// TIA Portal project "PolyMix_v0.1" (V14) (continued)
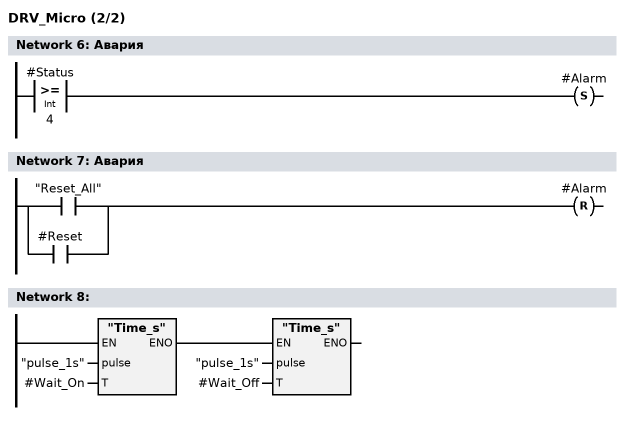
   RUNG wire#powerrail
      { S7_Templates := "SrcType := Int" } GE_Contact(in1 := #Status, in2 := 4)
      S_Coil( #Alarm )
   END_RUNG
   // the same network as SCL:
   IF #Status >= 4 THEN #Alarm := TRUE; END_IF;
END_REGION

REGION Network 7: Авария
   RUNG wire#powerrail
      Contact( "Reset_All" )
      wire#w1
      R_Coil( #Alarm )
   END_RUNG
   RUNG wire#powerrail
      Contact( #Reset )
   END_RUNG wire#w1
   // the same network as SCL:
   IF "Reset_All" OR #Reset THEN #Alarm := FALSE; END_IF;
END_REGION

REGION Network 8
   RUNG wire#powerrail
      "Time_s"(pulse := "pulse_1s", T := #Wait_On)
      "Time_s"(pulse := "pulse_1s", T := #Wait_Off)
   END_RUNG
   // the same network as SCL:
   "Time_s"(pulse := "pulse_1s", T := #Wait_On, ENO => #_w1);
   IF #_w1 THEN "Time_s"(pulse := "pulse_1s", T := #Wait_Off); END_IF;
END_REGION
END_FUNCTION_BLOCK

// folder: Modules

FUNCTION_BLOCK "DIx"   // FB200, LAD
{ S7_Optimized_Access := 'FALSE' }
VERSION : 0.1
// Input - входной сигнал контроллера
// pulse - частота фильтрации дребезга
// Signal - обработанный и отфильтрованный сигнал, используемый в дальнейшем
   VAR
      M1_FB_Ready : "DI_ex";   // I 0.0 - Мешалка 1 - готовность
      M1_FB_Run : "DI_ex";   // I 0.1 - Мешалка 1 - работа
      M2_FB_Ready : "DI_ex";   // I 0.2 - Мешалка 2 - готовность
      M2_FB_Run : "DI_ex";   // I 0.3 - Мешалка 2 - работа
      M3_FB_Ready : "DI_ex";   // I 0.4 - Мешалка 3 - готовность
      M3_FB_Run : "DI_ex";   // I 0.5 - Мешалка 3 - работа
      DD_FB_Ready : "DI_ex";   // I 0.6 - Дозатор сухого вещества - готовность
      Dos_FB_Run : "DI_ex";   // I 0.7 - Дозатор - работа
      DD_LLS : "DI_ex";   // I 1.0 - Дозатор сухого вещества - низкий уровень
      Vibro_FB_Ready : "DI_ex";   // I 1.1 - Вибратор - готовность
      Transporter : "DI_ex";   // I 1.2 - Пневмотранспортёр - готовность
      DL_FB_Ready : "DI_ex";   // I 1.3 - Дозатор жидкого вещества - готовность
      Dry_Run : "DI_ex";   // I 1.4 - Датчик протока
      AllBlock : "DI_ex";   // I 1.5 - Датчик перелива или Аварийная остановка
   END_VAR
   VAR_TEMP   // added for the SCL form of the ladder/FBD networks
      _w1 : Bool;
      _w2 : Bool;
   END_VAR
BEGIN

REGION Network 1: Мешалка 1
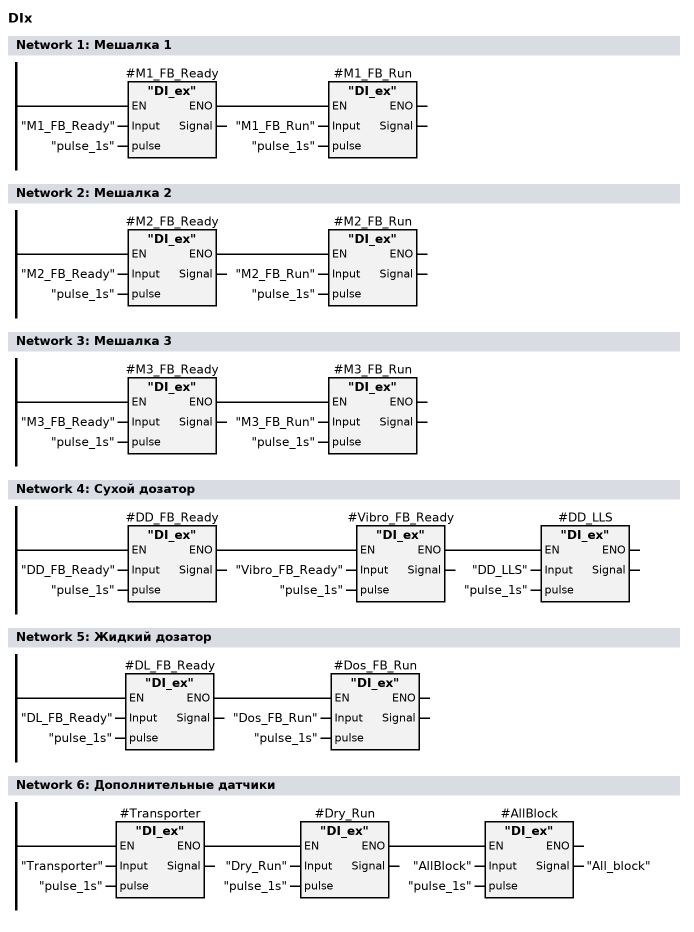
   RUNG wire#powerrail
      #M1_FB_Ready(Input := "M1_FB_Ready", pulse := "pulse_1s", Signal =>)
      #M1_FB_Run(Input := "M1_FB_Run", pulse := "pulse_1s", Signal =>)
   END_RUNG
   // the same network as SCL:
   #M1_FB_Ready(Input := "M1_FB_Ready", pulse := "pulse_1s", ENO => #_w1);   // "DI_ex"
   IF #_w1 THEN
       #M1_FB_Run(Input := "M1_FB_Run", pulse := "pulse_1s");   // "DI_ex"
   END_IF;
END_REGION

REGION Network 2: Мешалка 2
   RUNG wire#powerrail
      #M2_FB_Ready(Input := "M2_FB_Ready", pulse := "pulse_1s", Signal =>)
      #M2_FB_Run(Input := "M2_FB_Run", pulse := "pulse_1s", Signal =>)
   END_RUNG
   // the same network as SCL:
   #M2_FB_Ready(Input := "M2_FB_Ready", pulse := "pulse_1s", ENO => #_w1);   // "DI_ex"
   IF #_w1 THEN
       #M2_FB_Run(Input := "M2_FB_Run", pulse := "pulse_1s");   // "DI_ex"
   END_IF;
END_REGION

REGION Network 3: Мешалка 3
   RUNG wire#powerrail
      #M3_FB_Ready(Input := "M3_FB_Ready", pulse := "pulse_1s", Signal =>)
      #M3_FB_Run(Input := "M3_FB_Run", pulse := "pulse_1s", Signal =>)
   END_RUNG
   // the same network as SCL:
   #M3_FB_Ready(Input := "M3_FB_Ready", pulse := "pulse_1s", ENO => #_w1);   // "DI_ex"
   IF #_w1 THEN
       #M3_FB_Run(Input := "M3_FB_Run", pulse := "pulse_1s");   // "DI_ex"
   END_IF;
END_REGION

REGION Network 4: Сухой дозатор
   RUNG wire#powerrail
      #DD_FB_Ready(Input := "DD_FB_Ready", pulse := "pulse_1s", Signal =>)
      #Vibro_FB_Ready(Input := "Vibro_FB_Ready", pulse := "pulse_1s", Signal =>)
      #DD_LLS(Input := "DD_LLS", pulse := "pulse_1s", Signal =>)
   END_RUNG
   // the same network as SCL:
   #DD_FB_Ready(Input := "DD_FB_Ready", pulse := "pulse_1s", ENO => #_w1);   // "DI_ex"
   #Vibro_FB_Ready(EN := #_w1, Input := "Vibro_FB_Ready", pulse := "pulse_1s", ENO => #_w2);   // "DI_ex"
   IF #_w2 THEN
       #DD_LLS(Input := "DD_LLS", pulse := "pulse_1s");   // "DI_ex"
   END_IF;
END_REGION

REGION Network 5: Жидкий дозатор
   RUNG wire#powerrail
      #DL_FB_Ready(Input := "DL_FB_Ready", pulse := "pulse_1s", Signal =>)
      #Dos_FB_Run(Input := "Dos_FB_Run", pulse := "pulse_1s", Signal =>)
   END_RUNG
   // the same network as SCL:
   #DL_FB_Ready(Input := "DL_FB_Ready", pulse := "pulse_1s", ENO => #_w1);   // "DI_ex"
   IF #_w1 THEN
       #Dos_FB_Run(Input := "Dos_FB_Run", pulse := "pulse_1s");   // "DI_ex"
   END_IF;
END_REGION

REGION Network 6: Дополнительные датчики
   RUNG wire#powerrail
      #Transporter(Input := "Transporter", pulse := "pulse_1s", Signal =>)
      #Dry_Run(Input := "Dry_Run", pulse := "pulse_1s", Signal =>)
      #AllBlock(Input := "AllBlock", pulse := "pulse_1s", Signal => "All_block")
   END_RUNG
   // the same network as SCL:
   #Transporter(Input := "Transporter", pulse := "pulse_1s", ENO => #_w1);   // "DI_ex"
   #Dry_Run(EN := #_w1, Input := "Dry_Run", pulse := "pulse_1s", ENO => #_w2);   // "DI_ex"
   IF #_w2 THEN
       #AllBlock(Input := "AllBlock", pulse := "pulse_1s", Signal => "All_block");   // "DI_ex"
   END_IF;
END_REGION
END_FUNCTION_BLOCK

FUNCTION_BLOCK "DOx"   // FB201, LAD
{ S7_Optimized_Access := 'FALSE' }
VERSION : 0.1
// Start - управляющий сигнал из программы
// Q - выходной сигнал контроллера
// pulse - кратность времени в импульсном режиме
   VAR
      M1_CMD : "DO_ex";   // Q 0.0 - Мешалка 1 - запуск
      M2_CMD : "DO_ex";   // Q 0.1 - Мешалка 2 - запуск
      M3_CMD : "DO_ex";   // Q 0.2 - Мешалка 3 - запуск
      DD_CMD : "DO_ex";   // Q 0.3 - Дозатор сухого вещества - запуск
      Vibro_CMD : "DO_ex";   // Q 0.4 - Вибратор - запуск
      DL_CMD : "DO_ex";   // Q 0.5 - Дозатор жидкого вещества - запуск
      KC1_CMD : "DO_ex";   // Q 0.6 - Соленоидный клапан КС1
      LED_Dry_Run : "DO_ex";   // Q 0.7 - LED - сухой ход
      LED_Alarm : "DO_ex";   // Q 1.0 - LED - общая авария
      LED_Empty : "DO_ex";   // Q 1.1 - LED - бункер пуст
   END_VAR
   VAR_TEMP   // added for the SCL form of the ladder/FBD networks
      _w1 : Bool;
      _w2 : Bool;
   END_VAR
BEGIN

REGION Network 1: Мешалки 1-3
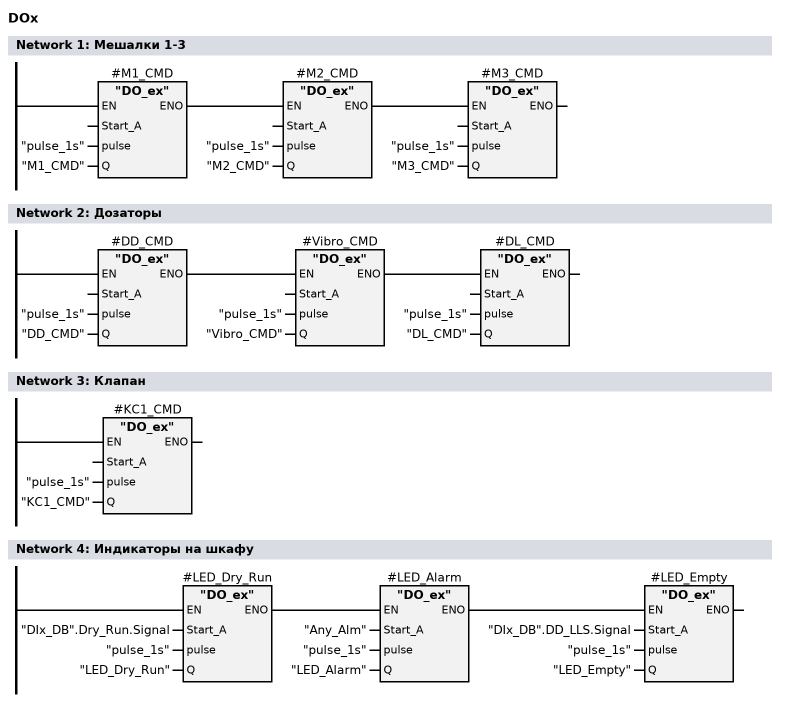
   RUNG wire#powerrail
      #M1_CMD(Start_A :=, pulse := "pulse_1s", Q := "M1_CMD")
      #M2_CMD(Start_A :=, pulse := "pulse_1s", Q := "M2_CMD")
      #M3_CMD(Start_A :=, pulse := "pulse_1s", Q := "M3_CMD")
   END_RUNG
   // the same network as SCL:
   #M1_CMD(pulse := "pulse_1s", Q := "M1_CMD", ENO => #_w1);   // "DO_ex"
   #M2_CMD(EN := #_w1, pulse := "pulse_1s", Q := "M2_CMD", ENO => #_w2);   // "DO_ex"
   IF #_w2 THEN
       #M3_CMD(pulse := "pulse_1s", Q := "M3_CMD");   // "DO_ex"
   END_IF;
END_REGION

REGION Network 2: Дозаторы
   RUNG wire#powerrail
      #DD_CMD(Start_A :=, pulse := "pulse_1s", Q := "DD_CMD")
      #Vibro_CMD(Start_A :=, pulse := "pulse_1s", Q := "Vibro_CMD")
      #DL_CMD(Start_A :=, pulse := "pulse_1s", Q := "DL_CMD")
   END_RUNG
   // the same network as SCL:
   #DD_CMD(pulse := "pulse_1s", Q := "DD_CMD", ENO => #_w1);   // "DO_ex"
   #Vibro_CMD(EN := #_w1, pulse := "pulse_1s", Q := "Vibro_CMD", ENO => #_w2);   // "DO_ex"
   IF #_w2 THEN
       #DL_CMD(pulse := "pulse_1s", Q := "DL_CMD");   // "DO_ex"
   END_IF;
END_REGION

REGION Network 3: Клапан
   RUNG wire#powerrail
      #KC1_CMD(Start_A :=, pulse := "pulse_1s", Q := "KC1_CMD")
   END_RUNG
   // the same network as SCL:
   #KC1_CMD(pulse := "pulse_1s", Q := "KC1_CMD");   // "DO_ex"
END_REGION

REGION Network 4: Индикаторы на шкафу
   RUNG wire#powerrail
      #LED_Dry_Run(Start_A := "DIx_DB".Dry_Run.Signal, pulse := "pulse_1s", Q := "LED_Dry_Run")
      #LED_Alarm(Start_A := "Any_Alm", pulse := "pulse_1s", Q := "LED_Alarm")
      #LED_Empty(Start_A := "DIx_DB".DD_LLS.Signal, pulse := "pulse_1s", Q := "LED_Empty")
   END_RUNG
   // the same network as SCL:
   #LED_Dry_Run(Start_A := "DIx_DB".Dry_Run.Signal, pulse := "pulse_1s", Q := "LED_Dry_Run", ENO => #_w1);   // "DO_ex"
   #LED_Alarm(EN := #_w1, Start_A := "Any_Alm", pulse := "pulse_1s", Q := "LED_Alarm", ENO => #_w2);   // "DO_ex"
   IF #_w2 THEN
       #LED_Empty(Start_A := "DIx_DB".DD_LLS.Signal, pulse := "pulse_1s", Q := "LED_Empty");   // "DO_ex"
   END_IF;
END_REGION
END_FUNCTION_BLOCK

FUNCTION_BLOCK "Micro"   // FB207, LAD
{ S7_Optimized_Access := 'FALSE' }
VERSION : 0.1
   VAR
      KC1 : "DRV_Micro";   // Соленоидный клапан
   END_VAR
   // KC1.No_FB := true;
BEGIN

REGION Network 1
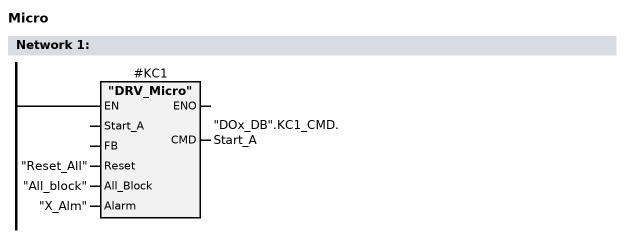
   RUNG wire#powerrail
      #KC1(Start_A :=, FB :=, Reset := "Reset_All", All_Block := "All_block", Alarm := "X_Alm", CMD => "DOx_DB".KC1_CMD.Start_A)
   END_RUNG
   // the same network as SCL:
   #KC1(Reset := "Reset_All", All_Block := "All_block", Alarm := "X_Alm", CMD => "DOx_DB".KC1_CMD.Start_A);   // "DRV_Micro"
END_REGION
END_FUNCTION_BLOCK

// folder: System

FUNCTION "DRV_pulse" : Void   // FC100, LAD
{ S7_Optimized_Access := 'FALSE' }
VERSION : 0.1
   VAR_TEMP   // added for the SCL form of the ladder/FBD networks
      _w1 : Bool;
      _w2 : Bool;
   END_VAR
BEGIN

REGION Network 1
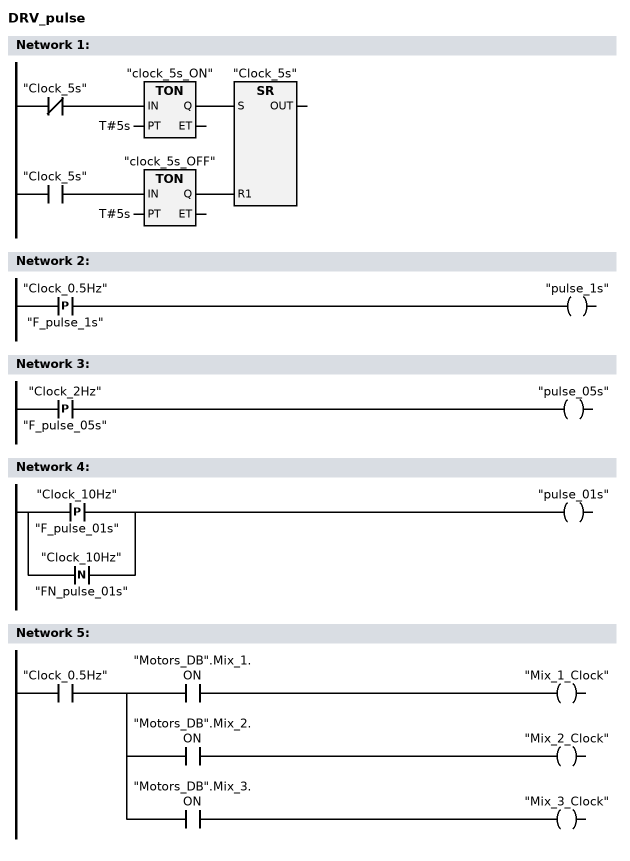
   "clock_5s_ON".TON(IN := NOT "Clock_5s", PT := T#5s);
   "clock_5s_OFF".TON(IN := "Clock_5s", PT := T#5s);
   IF "clock_5s_ON".Q THEN
       "Clock_5s" := TRUE;   // SR flip-flop
   END_IF;
   IF "clock_5s_OFF".Q THEN "Clock_5s" := FALSE; END_IF;
END_REGION

REGION Network 2
   RUNG wire#powerrail
      P_Contact(operand := "Clock_0.5Hz", bit := "F_pulse_1s")
      Coil( "pulse_1s" )
   END_RUNG
   // the same network as SCL:
   #_w1 := "Clock_0.5Hz" AND NOT "F_pulse_1s";   // rising edge of "Clock_0.5Hz"
   "F_pulse_1s" := "Clock_0.5Hz";
   "pulse_1s" := #_w1;
END_REGION

REGION Network 3
   RUNG wire#powerrail
      P_Contact(operand := "Clock_2Hz", bit := "F_pulse_05s")
      Coil( "pulse_05s" )
   END_RUNG
   // the same network as SCL:
   #_w1 := "Clock_2Hz" AND NOT "F_pulse_05s";   // rising edge of "Clock_2Hz"
   "F_pulse_05s" := "Clock_2Hz";
   "pulse_05s" := #_w1;
END_REGION

REGION Network 4
   RUNG wire#powerrail
      P_Contact(operand := "Clock_10Hz", bit := "F_pulse_01s")
      wire#w1
      Coil( "pulse_01s" )
   END_RUNG
   RUNG wire#powerrail
      N_Contact(operand := "Clock_10Hz", bit := "FN_pulse_01s")
   END_RUNG wire#w1
   // the same network as SCL:
   #_w1 := "Clock_10Hz" AND NOT "F_pulse_01s";   // rising edge of "Clock_10Hz"
   "F_pulse_01s" := "Clock_10Hz";
   #_w2 := NOT "Clock_10Hz" AND "FN_pulse_01s";   // falling edge of "Clock_10Hz"
   "FN_pulse_01s" := "Clock_10Hz";
   "pulse_01s" := #_w1 OR #_w2;
END_REGION

REGION Network 5
   RUNG wire#powerrail
      Contact( "Clock_0.5Hz" )
      wire#w1
      Contact( "Motors_DB".Mix_1.ON )
      Coil( "Mix_1_Clock" )
   END_RUNG
   RUNG wire#w1
      Contact( "Motors_DB".Mix_2.ON )
      Coil( "Mix_2_Clock" )
   END_RUNG
   RUNG wire#w1
      Contact( "Motors_DB".Mix_3.ON )
      Coil( "Mix_3_Clock" )
   END_RUNG
   // the same network as SCL:
   "Mix_1_Clock" := "Clock_0.5Hz" AND "Motors_DB".Mix_1.ON;
   "Mix_2_Clock" := "Clock_0.5Hz" AND "Motors_DB".Mix_2.ON;
   "Mix_3_Clock" := "Clock_0.5Hz" AND "Motors_DB".Mix_3.ON;
END_REGION
END_FUNCTION

FUNCTION "DRV_End" : Void   // FC101, LAD
{ S7_Optimized_Access := 'TRUE' }
VERSION : 0.1
BEGIN

REGION Network 1: Одно из устройств нижнего уровня в ручном режиме
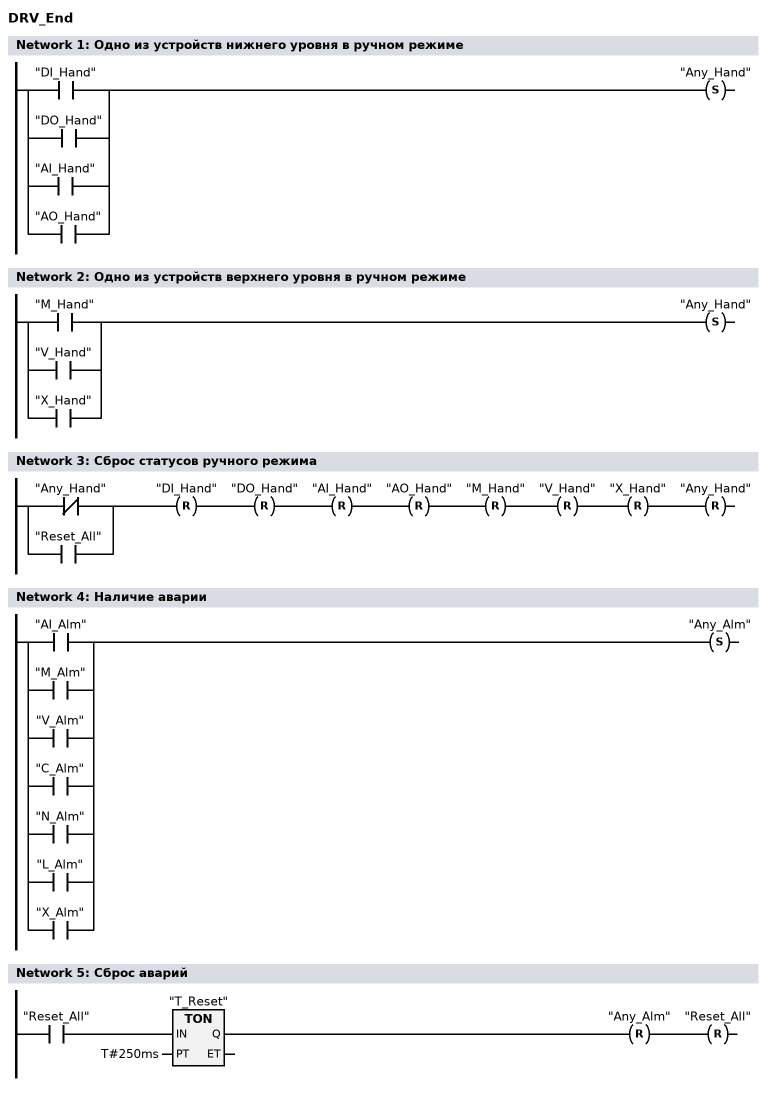
   RUNG wire#powerrail
      Contact( "DI_Hand" )
      wire#w1
      S_Coil( "Any_Hand" )
   END_RUNG
   RUNG wire#powerrail
      Contact( "DO_Hand" )
   END_RUNG wire#w1
   RUNG wire#powerrail
      Contact( "AI_Hand" )
   END_RUNG wire#w1
   RUNG wire#powerrail
      Contact( "AO_Hand" )
   END_RUNG wire#w1
   // the same network as SCL:
   IF "DI_Hand" OR "DO_Hand" OR "AI_Hand" OR "AO_Hand" THEN "Any_Hand" := TRUE; END_IF;
END_REGION

REGION Network 2: Одно из устройств верхнего уровня в ручном режиме
   RUNG wire#powerrail
      Contact( "M_Hand" )
      wire#w1
      S_Coil( "Any_Hand" )
   END_RUNG
   RUNG wire#powerrail
      Contact( "V_Hand" )
   END_RUNG wire#w1
   RUNG wire#powerrail
      Contact( "X_Hand" )
   END_RUNG wire#w1
   // the same network as SCL:
   IF "M_Hand" OR "V_Hand" OR "X_Hand" THEN "Any_Hand" := TRUE; END_IF;
END_REGION

REGION Network 3: Сброс статусов ручного режима
   RUNG wire#powerrail
      I_Contact( "Any_Hand" )
      wire#w1
      R_Coil( "DI_Hand" )
      R_Coil( "DO_Hand" )
      R_Coil( "AI_Hand" )
      R_Coil( "AO_Hand" )
      R_Coil( "M_Hand" )
      R_Coil( "V_Hand" )
      R_Coil( "X_Hand" )
      R_Coil( "Any_Hand" )
   END_RUNG
   RUNG wire#powerrail
      Contact( "Reset_All" )
   END_RUNG wire#w1
   // the same network as SCL:
   IF NOT "Any_Hand" OR "Reset_All" THEN
       "DI_Hand" := FALSE;
       "DO_Hand" := FALSE;
       "AI_Hand" := FALSE;
       "AO_Hand" := FALSE;
       "M_Hand" := FALSE;
       "V_Hand" := FALSE;
       "X_Hand" := FALSE;
       "Any_Hand" := FALSE;
   END_IF;
END_REGION

REGION Network 4: Наличие аварии
   RUNG wire#powerrail
      Contact( "AI_Alm" )
      wire#w1
      S_Coil( "Any_Alm" )
   END_RUNG
   RUNG wire#powerrail
      Contact( "M_Alm" )
   END_RUNG wire#w1
   RUNG wire#powerrail
      Contact( "V_Alm" )
   END_RUNG wire#w1
   RUNG wire#powerrail
      Contact( "C_Alm" )
   END_RUNG wire#w1
   RUNG wire#powerrail
      Contact( "N_Alm" )
   END_RUNG wire#w1
   RUNG wire#powerrail
      Contact( "L_Alm" )
   END_RUNG wire#w1
   RUNG wire#powerrail
      Contact( "X_Alm" )
   END_RUNG wire#w1
   // the same network as SCL:
   IF "AI_Alm" OR "M_Alm" OR "V_Alm" OR "C_Alm" OR "N_Alm" OR "L_Alm" OR "X_Alm" THEN
       "Any_Alm" := TRUE;
   END_IF;
END_REGION

REGION Network 5: Сброс аварий
   "T_Reset".TON(IN := "Reset_All", PT := T#250ms);
   IF "T_Reset".Q THEN
       "Any_Alm" := FALSE;
       "Reset_All" := FALSE;
   END_IF;
END_REGION
END_FUNCTION

FUNCTION "Converter" : Void   // FC102, LAD
TITLE = Драйвер линеаризации аналогового сигнала
{ S7_Optimized_Access := 'FALSE' }
VERSION : 0.1
   VAR_INPUT
      Converter : Struct
         Use_Min_In : Bool;   // Отсекать входные значения ниже минимума
         Use_Max_In : Bool;   // Отсекать входные значения выше максимума
         Use_Min_Out : Bool;   // Отсекать результат ниже минимума
         Use_Max_Out : Bool;   // Отсекать результат выше максимума
         Min_In : Real;   // Минимальный входной сигнал
         Max_In : Real;   // Максимальный входной сигнал
         Min_Out : Real;   // Минимальный выходной сигнал
         Max_Out : Real;   // Максимальный выходной сигнал
      END_STRUCT;
   END_VAR
   VAR_IN_OUT
      Signal : Real;   // Входной сигнал
      Result : Real;   // Результат линеаризации
   END_VAR
   VAR_TEMP
      Range_In : Real;   // Диапазон входного сигнала
      Range_Out : Real;   // Диапазон выходного сигнала
      T_T : Real;   // Соотношение диапазонов
      R_Sig : Real;   // Поправка на отрицательные значения
   END_VAR
BEGIN

REGION Network 1: Проверка нижнего уровня входного сигнала
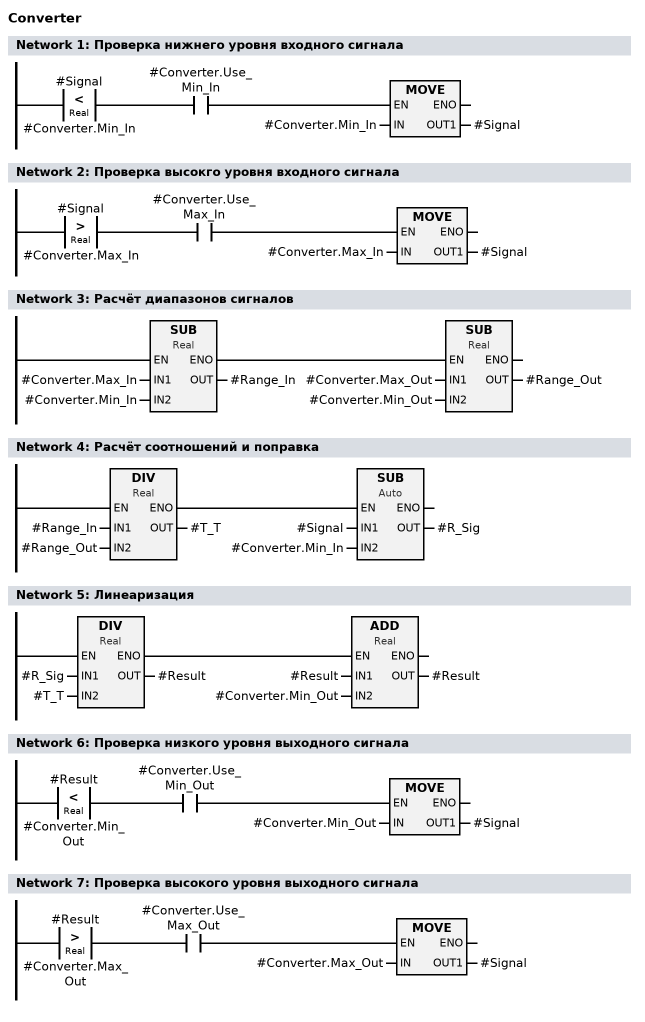
   RUNG wire#powerrail
      { S7_Templates := "SrcType := Real" } LT_Contact(in1 := #Signal, in2 := #Converter.Min_In)
      Contact( #Converter.Use_Min_In )
      Move(in := #Converter.Min_In, out1 => #Signal)
   END_RUNG
   // the same network as SCL:
   IF (#Signal < #Converter.Min_In) AND #Converter.Use_Min_In THEN #Signal := #Converter.Min_In; END_IF;
END_REGION

REGION Network 2: Проверка высокго уровня входного сигнала
   RUNG wire#powerrail
      { S7_Templates := "SrcType := Real" } GT_Contact(in1 := #Signal, in2 := #Converter.Max_In)
      Contact( #Converter.Use_Max_In )
      Move(in := #Converter.Max_In, out1 => #Signal)
   END_RUNG
   // the same network as SCL:
   IF (#Signal > #Converter.Max_In) AND #Converter.Use_Max_In THEN #Signal := #Converter.Max_In; END_IF;
END_REGION

REGION Network 3: Расчёт диапазонов сигналов
   RUNG wire#powerrail
      { S7_Templates := "SrcType := Real"; S7_GenerateENO := "TRUE" } Sub(in1 := #Converter.Max_In, in2 := #Converter.Min_In, out => #Range_In)
      { S7_Templates := "SrcType := Real"; S7_GenerateENO := "TRUE" } Sub(in1 := #Converter.Max_Out, in2 := #Converter.Min_Out, out => #Range_Out)
   END_RUNG
   // the same network as SCL:
   // ENO of a box is taken as its EN; it also drops when the box reports an error
   #Range_In := #Converter.Max_In - #Converter.Min_In;
   #Range_Out := #Converter.Max_Out - #Converter.Min_Out;
END_REGION

REGION Network 4: Расчёт соотношений и поправка
   RUNG wire#powerrail
      { S7_Templates := "SrcType := Real"; S7_GenerateENO := "TRUE" } Div(in1 := #Range_In, in2 := #Range_Out, out => #T_T)
      Sub(in1 := #Signal, in2 := #Converter.Min_In, out => #R_Sig)
   END_RUNG
   // the same network as SCL:
   // ENO of a box is taken as its EN; it also drops when the box reports an error
   #T_T := #Range_In / #Range_Out;
   #R_Sig := #Signal - #Converter.Min_In;
END_REGION

REGION Network 5: Линеаризация
   RUNG wire#powerrail
      { S7_Templates := "SrcType := Real"; S7_GenerateENO := "TRUE" } Div(in1 := #R_Sig, in2 := #T_T, out => #Result)
      { S7_Templates := "SrcType := Real"; S7_GenerateENO := "TRUE" } Add(in1 := #Result, in2 := #Converter.Min_Out, out => #Result)
   END_RUNG
   // the same network as SCL:
   // ENO of a box is taken as its EN; it also drops when the box reports an error
   #Result := #R_Sig / #T_T;
   #Result := #Result + #Converter.Min_Out;
END_REGION

REGION Network 6: Проверка низкого уровня выходного сигнала
   RUNG wire#powerrail
      { S7_Templates := "SrcType := Real" } LT_Contact(in1 := #Result, in2 := #Converter.Min_Out)
      Contact( #Converter.Use_Min_Out )
      Move(in := #Converter.Min_Out, out1 => #Signal)
   END_RUNG
   // the same network as SCL:
   IF (#Result < #Converter.Min_Out) AND #Converter.Use_Min_Out THEN #Signal := #Converter.Min_Out; END_IF;
END_REGION

REGION Network 7: Проверка высокого уровня выходного сигнала
   RUNG wire#powerrail
      { S7_Templates := "SrcType := Real" } GT_Contact(in1 := #Result, in2 := #Converter.Max_Out)
      Contact( #Converter.Use_Max_Out )
      Move(in := #Converter.Max_Out, out1 => #Signal)
   END_RUNG
   // the same network as SCL:
   IF (#Result > #Converter.Max_Out) AND #Converter.Use_Max_Out THEN #Signal := #Converter.Max_Out; END_IF;
END_REGION
END_FUNCTION

FUNCTION "INV" : Void   // FC111, LAD
{ S7_Optimized_Access := 'TRUE' }
VERSION : 0.1
   VAR_INPUT
      S : Bool;   // Сигнал
      I : Bool;   // Инверсия
   END_VAR
   VAR_IN_OUT
      R : Bool;   // Результат
   END_VAR
BEGIN

REGION Network 1: Инверсия сигнала
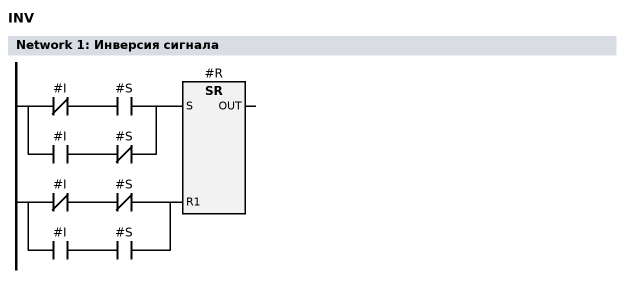
   RUNG wire#powerrail
      I_Contact( #I )
      Contact( #S )
      wire#w1
      S_SR(operand := #R, r1 := wire#w2)
   END_RUNG
   RUNG wire#powerrail
      Contact( #I )
      I_Contact( #S )
   END_RUNG wire#w1
   RUNG wire#powerrail
      I_Contact( #I )
      I_Contact( #S )
   END_RUNG wire#w2
   RUNG wire#powerrail
      Contact( #I )
      Contact( #S )
   END_RUNG wire#w2
   // the same network as SCL:
   IF (NOT #I AND #S) OR (#I AND NOT #S) THEN
       #R := TRUE;   // SR flip-flop
   END_IF;
   IF (NOT #I AND NOT #S) OR (#I AND #S) THEN #R := FALSE; END_IF;
END_REGION
END_FUNCTION

FUNCTION "Mode" : Void   // FC150, LAD
{ S7_Optimized_Access := 'FALSE' }
VERSION : 0.1
   VAR_INPUT
      CMD : Struct   // Основные команды
         Hand : Bool;   // 0 - авто, 1 - ручной / 0 - Авто, 1 - Ручной
         Start_A : Bool;   // Автозапуск / Запуск в авторежиме
         Start_M : Bool;   // Ручной - вперёд / Запуск в ручном режиме
         Force : Bool;   // Принудительный
         Lock : Bool;   // Блокировать / Блокировка
         Local : Bool;   // Локальный
         Service : Bool;   // Сервис
         Safety : Bool;   // Безопасность
         Alarm : Bool;   // Есть авария / Авария
         Reset : Bool;   // Сброс аварий
         Sim : Bool;   // Режим симуляции
      END_STRUCT;
      All_Block : Bool;   // Аварийная блокировка
   END_VAR
   VAR_OUTPUT
      Mode : Int;   // Режим работы
   END_VAR
BEGIN

REGION Network 1: Автоматический режим
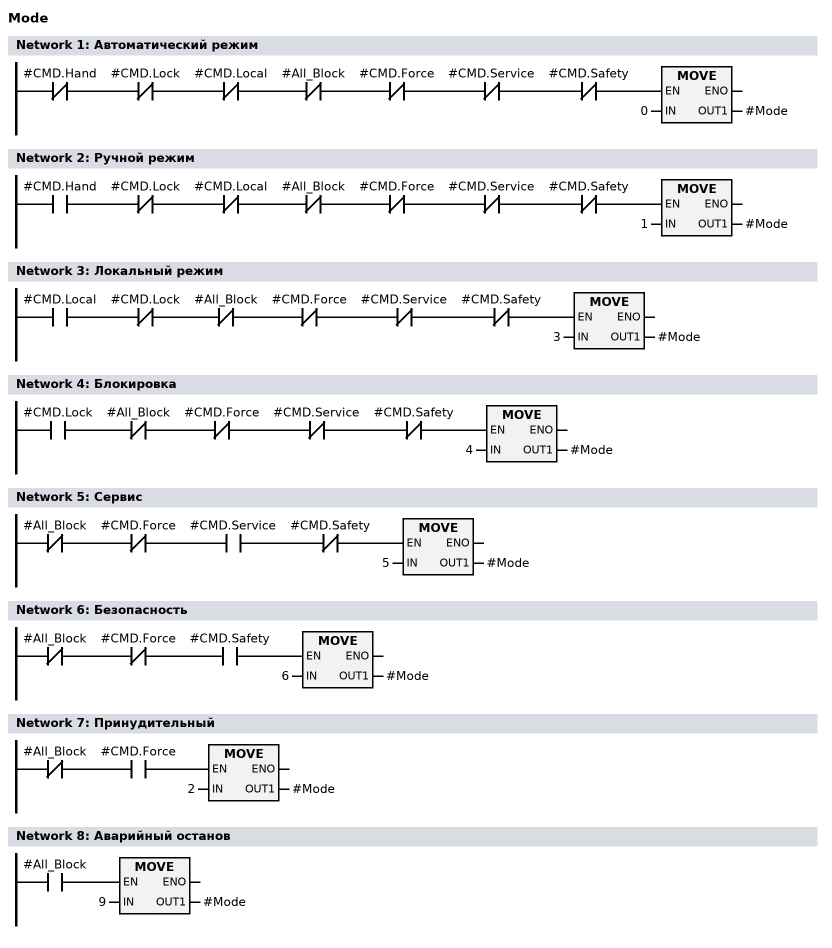
   RUNG wire#powerrail
      I_Contact( #CMD.Hand )
      I_Contact( #CMD.Lock )
      I_Contact( #CMD.Local )
      I_Contact( #All_Block )
      I_Contact( #CMD.Force )
      I_Contact( #CMD.Service )
      I_Contact( #CMD.Safety )
      { S7_GenerateENO := "TRUE" } Move(in := 0, out1 => #Mode)
   END_RUNG
   // the same network as SCL:
   IF NOT #CMD.Hand AND NOT #CMD.Lock AND NOT #CMD.Local AND NOT #All_Block AND NOT #CMD.Force AND NOT #CMD.Service AND NOT #CMD.Safety THEN
       #Mode := 0;
   END_IF;
END_REGION

REGION Network 2: Ручной режим
   RUNG wire#powerrail
      Contact( #CMD.Hand )
      I_Contact( #CMD.Lock )
      I_Contact( #CMD.Local )
      I_Contact( #All_Block )
      I_Contact( #CMD.Force )
      I_Contact( #CMD.Service )
      I_Contact( #CMD.Safety )
      { S7_GenerateENO := "TRUE" } Move(in := 1, out1 => #Mode)
   END_RUNG
   // the same network as SCL:
   IF #CMD.Hand AND NOT #CMD.Lock AND NOT #CMD.Local AND NOT #All_Block AND NOT #CMD.Force AND NOT #CMD.Service AND NOT #CMD.Safety THEN
       #Mode := 1;
   END_IF;
END_REGION

REGION Network 3: Локальный режим
   RUNG wire#powerrail
      Contact( #CMD.Local )
      I_Contact( #CMD.Lock )
      I_Contact( #All_Block )
      I_Contact( #CMD.Force )
      I_Contact( #CMD.Service )
      I_Contact( #CMD.Safety )
      { S7_GenerateENO := "TRUE" } Move(in := 3, out1 => #Mode)
   END_RUNG
   // the same network as SCL:
   IF #CMD.Local AND NOT #CMD.Lock AND NOT #All_Block AND NOT #CMD.Force AND NOT #CMD.Service AND NOT #CMD.Safety THEN
       #Mode := 3;
   END_IF;
END_REGION

REGION Network 4: Блокировка
   RUNG wire#powerrail
      Contact( #CMD.Lock )
      I_Contact( #All_Block )
      I_Contact( #CMD.Force )
      I_Contact( #CMD.Service )
      I_Contact( #CMD.Safety )
      { S7_GenerateENO := "TRUE" } Move(in := 4, out1 => #Mode)
   END_RUNG
   // the same network as SCL:
   IF #CMD.Lock AND NOT #All_Block AND NOT #CMD.Force AND NOT #CMD.Service AND NOT #CMD.Safety THEN
       #Mode := 4;
   END_IF;
END_REGION

REGION Network 5: Сервис
   RUNG wire#powerrail
      I_Contact( #All_Block )
      I_Contact( #CMD.Force )
      Contact( #CMD.Service )
      I_Contact( #CMD.Safety )
      { S7_GenerateENO := "TRUE" } Move(in := 5, out1 => #Mode)
   END_RUNG
   // the same network as SCL:
   IF NOT #All_Block AND NOT #CMD.Force AND #CMD.Service AND NOT #CMD.Safety THEN #Mode := 5; END_IF;
END_REGION

REGION Network 6: Безопасность
   RUNG wire#powerrail
      I_Contact( #All_Block )
      I_Contact( #CMD.Force )
      Contact( #CMD.Safety )
      { S7_GenerateENO := "TRUE" } Move(in := 6, out1 => #Mode)
   END_RUNG
   // the same network as SCL:
   IF NOT #All_Block AND NOT #CMD.Force AND #CMD.Safety THEN #Mode := 6; END_IF;
END_REGION

REGION Network 7: Принудительный
   RUNG wire#powerrail
      I_Contact( #All_Block )
      Contact( #CMD.Force )
      { S7_GenerateENO := "TRUE" } Move(in := 2, out1 => #Mode)
   END_RUNG
   // the same network as SCL:
   IF NOT #All_Block AND #CMD.Force THEN #Mode := 2; END_IF;
END_REGION

REGION Network 8: Аварийный останов
   RUNG wire#powerrail
      Contact( #All_Block )
      { S7_GenerateENO := "TRUE" } Move(in := 9, out1 => #Mode)
   END_RUNG
   // the same network as SCL:
   IF #All_Block THEN #Mode := 9; END_IF;
END_REGION
END_FUNCTION

// ===== PLC "PLC_Master"  CPU 1214C DC/DC/DC =====
// protected blocks, not shown: "AI_ex", "AIx", "AO_ex", "AOx", "DRV_M_D", "Logick", "Motors", "PLF_FC", "Ponts", "RS232", "Statistics", "Time_m", "Time_r", "Time_s"

VAR_GLOBAL   // PLC tag table "Default tag table"
   "Sync_1" AT %M10.0 : Bool;
   "Sync_2" AT %M10.1 : Bool;
END_VAR

VAR_GLOBAL   // PLC tag table "IO"
   "M1_QF" AT %I0.0 : Bool;
   "M1_CMD" AT %Q0.0 : Bool;
   "LED_M1_Alarm" AT %Q0.6 : Bool;
   "M1_SP" AT %QW256 : Int;
   "M2_QF" AT %I0.1 : Bool;
   "M2_CMD" AT %Q0.1 : Bool;
   "LED_M2_Alarm" AT %Q0.7 : Bool;
   "M2_SP" AT %QW258 : Int;
   "M3_QF" AT %I0.2 : Bool;
   "M3_CMD" AT %Q0.2 : Bool;
   "LED_M3_Alarm" AT %Q1.0 : Bool;
   "M3_SP" AT %QW260 : Int;
   "Flow_1" AT %IW260 : Int;
   "Flow_2" AT %IW262 : Int;
   "Heat_1_Run" AT %I0.3 : Bool;
   "Heat_2_Run" AT %I0.4 : Bool;
   "Heat_3_Run" AT %I0.5 : Bool;
   "Heat_4_Run" AT %I0.6 : Bool;
   "Trans_1" AT %IW264 : Int;
   "Trans_2" AT %IW266 : Int;
   "AllBlock" AT %I0.7 : Bool;
   "Mass_1_Ready" AT %I1.0 : Bool;
   "Mass_2_Ready" AT %I1.1 : Bool;
   "LED_Error_1" AT %Q0.3 : Bool;
   "LED_Error_2" AT %Q0.4 : Bool;
   "LED_Alarm" AT %Q0.5 : Bool;
   "Flow_3" AT %IW268 : Int;
   "Flow_4" AT %IW270 : Int;
END_VAR

VAR_GLOBAL   // PLC tag table "Sys"
   "pulse_01s" AT %M2.0 : Bool;
   "pulse_05s" AT %M2.1 : Bool;
   "pulse_1s" AT %M2.2 : Bool;
   "All_block" AT %M3.0 : Bool;
   "Reset_All" AT %M3.1 : Bool;
   "Sim_All" AT %M3.2 : Bool;
   "Any_Hand" AT %M5.0 : Bool;
   "DI_Hand" AT %M5.1 : Bool;
   "DO_Hand" AT %M5.2 : Bool;
   "AI_Hand" AT %M5.3 : Bool;
   "AO_Hand" AT %M5.4 : Bool;
   "M_Hand" AT %M5.5 : Bool;
   "V_Hand" AT %M5.6 : Bool;
   "X_Hand" AT %M5.7 : Bool;
   "System_Byte" AT %MB1 : Byte;
   "FirstScan" AT %M1.0 : Bool;
   "DiagStatusUpdate" AT %M1.1 : Bool;
   "ON" AT %M1.2 : Bool;
   "OFF" AT %M1.3 : Bool;
   "Clock_Byte" AT %MB0 : Byte;
   "Clock_10Hz" AT %M0.0 : Bool;
   "Clock_5Hz" AT %M0.1 : Bool;
   "Clock_2.5Hz" AT %M0.2 : Bool;
   "Clock_2Hz" AT %M0.3 : Bool;
   "Clock_1.25Hz" AT %M0.4 : Bool;
   "Clock_1Hz" AT %M0.5 : Bool;
   "Clock_0.625Hz" AT %M0.6 : Bool;
   "Clock_0.5Hz" AT %M0.7 : Bool;
   "F_pulse_01s" AT %M2.3 : Bool;
   "F_pulse_05s" AT %M2.4 : Bool;
   "F_pulse_1s" AT %M2.5 : Bool;
   "FN_pulse_01s" AT %M2.6 : Bool;
   "Clock_5s" AT %M2.7 : Bool;
   "Any_Alm" AT %M6.0 : Bool;
   "AI_Alm" AT %M6.1 : Bool;
   "M_Alm" AT %M6.2 : Bool;
   "V_Alm" AT %M6.3 : Bool;
   "C_Alm" AT %M6.4 : Bool;
   "N_Alm" AT %M6.5 : Bool;
   "L_Alm" AT %M6.6 : Bool;
   "X_Alm" AT %M6.7 : Bool;
END_VAR

DATA_BLOCK "PID_M1"   // DB5
{ S7_Optimized_Access := 'FALSE' }
VERSION : 0.1
// stored: InstanceOfName PID_ex
"PID_ex"
BEGIN
   SP_P := 0.75;
   Max_SP := 2000.0;
   Max_in := 2500.0;
   Max_out := 1.3;
   Min_out := 0.7;
END_DATA_BLOCK

DATA_BLOCK "PID_M2"   // DB6
{ S7_Optimized_Access := 'FALSE' }
VERSION : 0.1
// stored: InstanceOfName PID_ex
"PID_ex"
BEGIN
   SP_P := 0.75;
   Max_SP := 2000.0;
   Max_in := 2500.0;
   Max_out := 1.3;
   Min_out := 0.7;
END_DATA_BLOCK

DATA_BLOCK "Comm_1_DB"   // DB11
{ S7_Optimized_Access := 'FALSE' }
VERSION : 0.1
   VAR
      DD_Status : Int;
      DD_Mode : Int;
      DD_Alarm : Word;
      DL_Status : Int;
      DL_Mode : Int;
      DL_Alarm : Word;
      Mix_1_Status : Int;
      Mix_1_Mode : Int;
      Mix_1_Alarm : Word;
      Mix_2_Status : Int;
      Mix_2_Mode : Int;
      Mix_2_Alarm : Word;
      Mix_3_Status : Int;
      Mix_3_Mode : Int;
      Mix_3_Alarm : Word;
      KC1_Status : Int;
      Flowmeter : Real;
      Flow_Alarm : Word;
      Level : Real;
      Level_Alarm : Word;
      SP : Real;
      Start : Bool;
      Hand : Bool;
      Warning : Bool;
      Config : Struct
         Use_DD : Bool;   // Использовать сухой дозатор
         Use_DL : Bool;   // Использовать жидкий дозатор
         Use_Mix_1 : Bool;   // Использовать мешалку 1
         Use_Mix_2 : Bool;   // Использовать мешалку 2
         Use_Mix_3 : Bool;   // Использовать мешалку 3
      END_STRUCT;
      Alarm : Word;
   END_VAR
BEGIN
END_DATA_BLOCK

DATA_BLOCK "Comm_2_DB"   // DB12
{ S7_Optimized_Access := 'FALSE' }